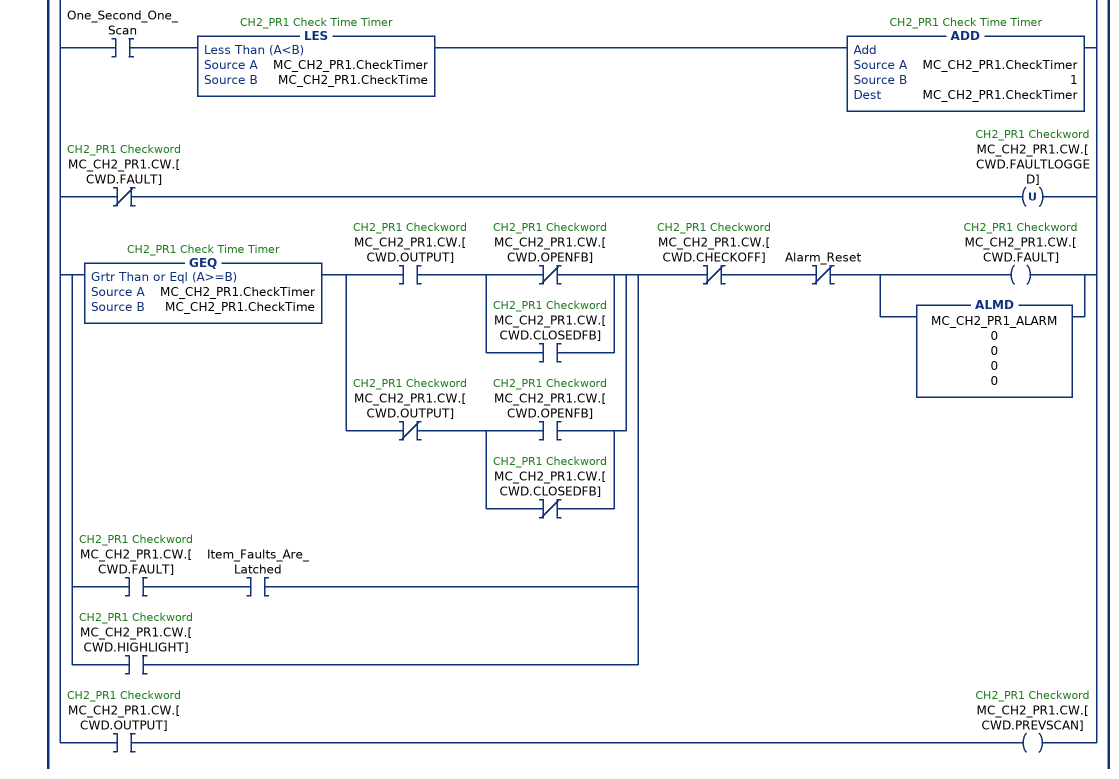
   38: [NEQ(MC_CH2_PR1.DriveBits,0) OTE(MC_CH2_PR1.CW.[CWD.AUTODRV]) ,[XIC(MC_CH2_PR1.CW.[CWD.AUTODRV]) XIO(MC_CH2_PR1.CW.[CWD.MANUAL]) ,XIC(MC_CH2_PR1.CW.[CWD.MANDRV]) XIC(MC_CH2_PR1.CW.[CWD.MANUAL]) ] OTE(MC_CH2_PR1.CW.[CWD.OUTPUT]) ,XIC(MC_CH2_PR1.CW.[CWD.OUTPUT]) OTE(MC_CH2_PR1_DR) ,XIC(S:FS) [OTU(MC_CH2_PR1.CW.[CWD.MANUAL]) ,LEQ(MC_CH2_PR1.CheckTime,0) MOV(Default_Check_Time,MC_CH2_PR1.CheckTime) ] ,[[XIC(MC_CH2_PR1_O) XIO(Item_Simulation_Flag) ,XIC(Item_Simulation_Flag) XIC(MC_CH2_PR1.CW.[CWD.OUTPUT]) XIO(MC_CH2_PR1.CW.[CWD.SIMFAIL]) ] OTE(MC_CH2_PR1.CW.[CWD.OPENFB]) ,[XIC(MC_CH2_PR1_C) XIO(Item_Simulation_Flag) ,XIC(Item_Simulation_Flag) XIO(MC_CH2_PR1.CW.[CWD.OUTPUT]) XIO(MC_CH2_PR1.CW.[CWD.SIMFAIL]) ] OTE(MC_CH2_PR1.CW.[CWD.CLOSEDFB]) ] ,[XIC(MC_CH2_PR1.CW.[CWD.OUTPUT]) XIO(MC_CH2_PR1.CW.[CWD.PREVSCAN]) ,XIO(MC_CH2_PR1.CW.[CWD.OUTPUT]) XIC(MC_CH2_PR1.CW.[CWD.PREVSCAN]) ] CLR(MC_CH2_PR1.CheckTimer) ,XIC(One_Second_One_Scan) LES(MC_CH2_PR1.CheckTimer,MC_CH2_PR1.CheckTime) ADD(MC_CH2_PR1.CheckTimer,1,MC_CH2_PR1.CheckTimer) ,XIO(MC_CH2_PR1.CW.[CWD.FAULT]) OTU(MC_CH2_PR1.CW.[CWD.FAULTLOGGED]) ,[GEQ(MC_CH2_PR1.CheckTimer,MC_CH2_PR1.CheckTime) [XIC(MC_CH2_PR1.CW.[CWD.OUTPUT]) [XIO(MC_CH2_PR1.CW.[CWD.OPENFB]) ,XIC(MC_CH2_PR1.CW.[CWD.CLOSEDFB]) ] ,XIO(MC_CH2_PR1.CW.[CWD.OUTPUT]) [XIC(MC_CH2_PR1.CW.[CWD.OPENFB]) ,XIO(MC_CH2_PR1.CW.[CWD.CLOSEDFB]) ] ] ,XIC(MC_CH2_PR1.CW.[CWD.FAULT]) XIC(Item_Faults_Are_Latched) ,XIC(MC_CH2_PR1.CW.[CWD.HIGHLIGHT]) ] XIO(MC_CH2_PR1.CW.[CWD.CHECKOFF]) XIO(Alarm_Reset) [OTE(MC_CH2_PR1.CW.[CWD.FAULT]) ,ALMD(MC_CH2_PR1_ALARM,0,0,0,0) ] ,XIC(MC_CH2_PR1.CW.[CWD.OUTPUT]) OTE(MC_CH2_PR1.CW.[CWD.PREVSCAN]) ];
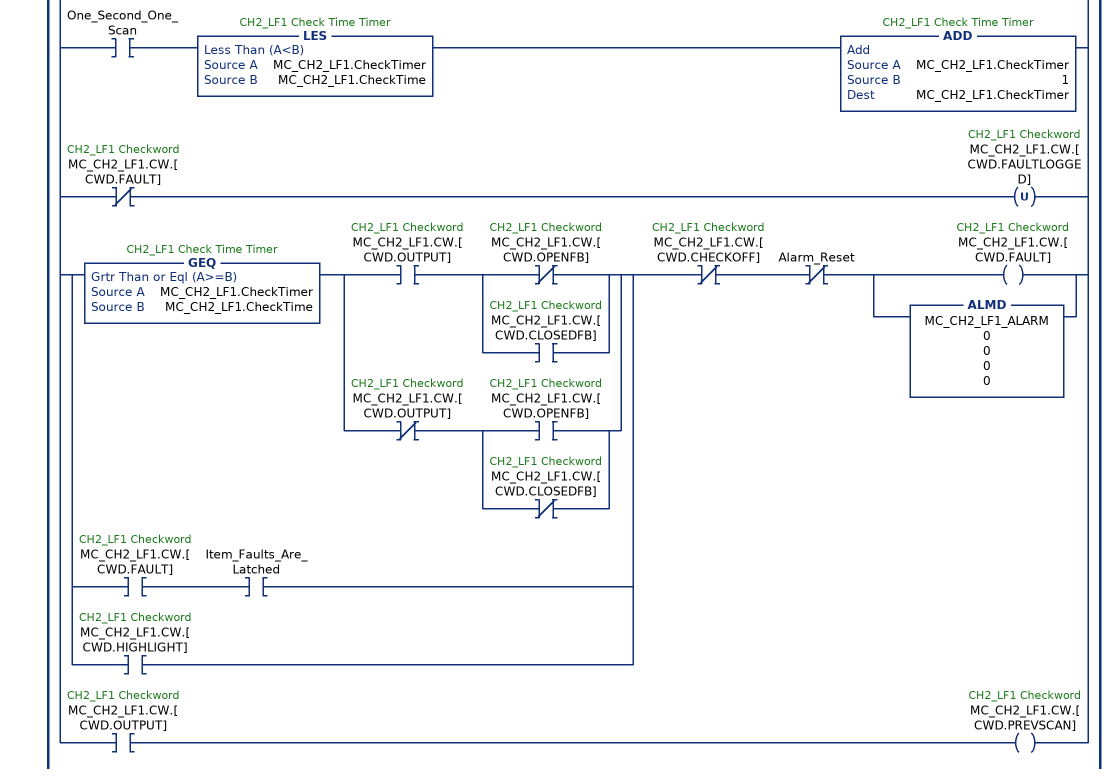
   39: [NEQ(MC_CH2_LF1.DriveBits,0) OTE(MC_CH2_LF1.CW.[CWD.AUTODRV]) ,[XIC(MC_CH2_LF1.CW.[CWD.AUTODRV]) XIO(MC_CH2_LF1.CW.[CWD.MANUAL]) ,XIC(MC_CH2_LF1.CW.[CWD.MANDRV]) XIC(MC_CH2_LF1.CW.[CWD.MANUAL]) ] OTE(MC_CH2_LF1.CW.[CWD.OUTPUT]) ,XIC(MC_CH2_LF1.CW.[CWD.OUTPUT]) OTE(MC_CH2_LF1_DR) ,XIC(S:FS) [OTU(MC_CH2_LF1.CW.[CWD.MANUAL]) ,LEQ(MC_CH2_LF1.CheckTime,0) MOV(Default_Check_Time,MC_CH2_LF1.CheckTime) ] ,[[XIC(MC_CH2_LF1_O) XIO(Item_Simulation_Flag) ,XIC(Item_Simulation_Flag) XIC(MC_CH2_LF1.CW.[CWD.OUTPUT]) XIO(MC_CH2_LF1.CW.[CWD.SIMFAIL]) ] OTE(MC_CH2_LF1.CW.[CWD.OPENFB]) ,[XIC(MC_CH2_LF1_C) XIO(Item_Simulation_Flag) ,XIC(Item_Simulation_Flag) XIO(MC_CH2_LF1.CW.[CWD.OUTPUT]) XIO(MC_CH2_LF1.CW.[CWD.SIMFAIL]) ] OTE(MC_CH2_LF1.CW.[CWD.CLOSEDFB]) ] ,[XIC(MC_CH2_LF1.CW.[CWD.OUTPUT]) XIO(MC_CH2_LF1.CW.[CWD.PREVSCAN]) ,XIO(MC_CH2_LF1.CW.[CWD.OUTPUT]) XIC(MC_CH2_LF1.CW.[CWD.PREVSCAN]) ] CLR(MC_CH2_LF1.CheckTimer) ,XIC(One_Second_One_Scan) LES(MC_CH2_LF1.CheckTimer,MC_CH2_LF1.CheckTime) ADD(MC_CH2_LF1.CheckTimer,1,MC_CH2_LF1.CheckTimer) ,XIO(MC_CH2_LF1.CW.[CWD.FAULT]) OTU(MC_CH2_LF1.CW.[CWD.FAULTLOGGED]) ,[GEQ(MC_CH2_LF1.CheckTimer,MC_CH2_LF1.CheckTime) [XIC(MC_CH2_LF1.CW.[CWD.OUTPUT]) [XIO(MC_CH2_LF1.CW.[CWD.OPENFB]) ,XIC(MC_CH2_LF1.CW.[CWD.CLOSEDFB]) ] ,XIO(MC_CH2_LF1.CW.[CWD.OUTPUT]) [XIC(MC_CH2_LF1.CW.[CWD.OPENFB]) ,XIO(MC_CH2_LF1.CW.[CWD.CLOSEDFB]) ] ] ,XIC(MC_CH2_LF1.CW.[CWD.FAULT]) XIC(Item_Faults_Are_Latched) ,XIC(MC_CH2_LF1.CW.[CWD.HIGHLIGHT]) ] XIO(MC_CH2_LF1.CW.[CWD.CHECKOFF]) XIO(Alarm_Reset) [OTE(MC_CH2_LF1.CW.[CWD.FAULT]) ,ALMD(MC_CH2_LF1_ALARM,0,0,0,0) ] ,XIC(MC_CH2_LF1.CW.[CWD.OUTPUT]) OTE(MC_CH2_LF1.CW.[CWD.PREVSCAN]) ];
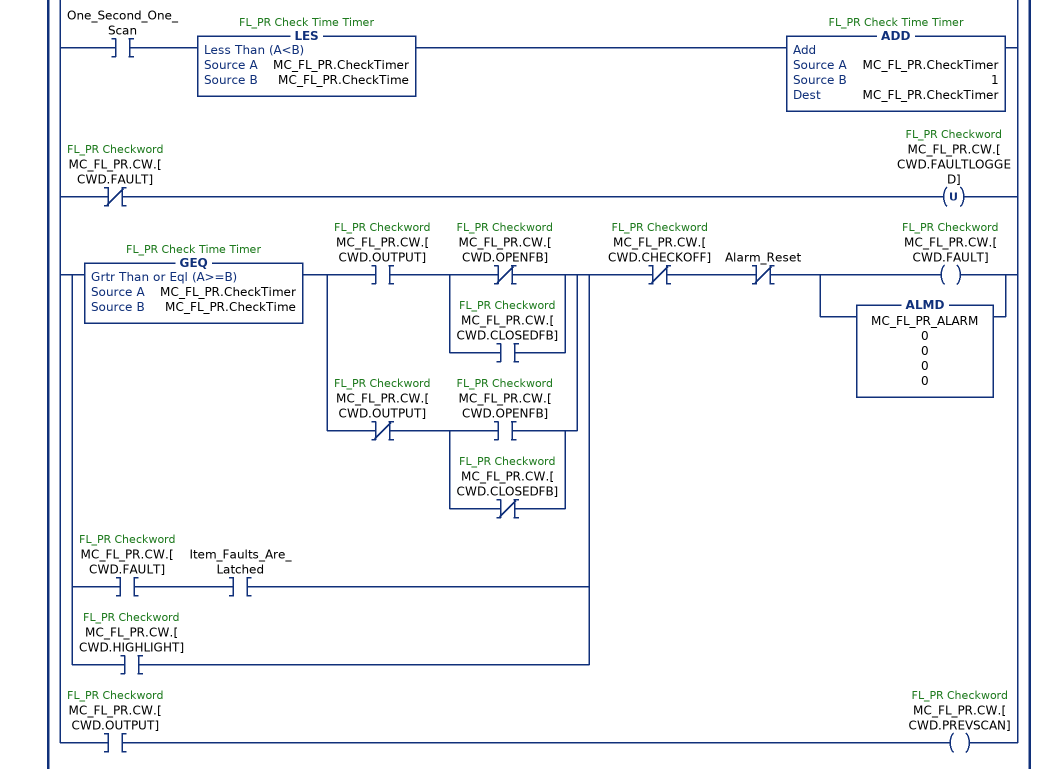
   40: [NEQ(MC_FL_PR.DriveBits,0) OTE(MC_FL_PR.CW.[CWD.AUTODRV]) ,[XIC(MC_FL_PR.CW.[CWD.AUTODRV]) XIO(MC_FL_PR.CW.[CWD.MANUAL]) ,XIC(MC_FL_PR.CW.[CWD.MANDRV]) XIC(MC_FL_PR.CW.[CWD.MANUAL]) ] OTE(MC_FL_PR.CW.[CWD.OUTPUT]) ,XIC(MC_FL_PR.CW.[CWD.OUTPUT]) OTE(MC_FL_PR_DR) ,XIC(S:FS) [OTU(MC_FL_PR.CW.[CWD.MANUAL]) ,LEQ(MC_FL_PR.CheckTime,0) MOV(Default_Check_Time,MC_FL_PR.CheckTime) ] ,[[XIC(MC_FL_PR_O) XIO(Item_Simulation_Flag) ,XIC(Item_Simulation_Flag) XIC(MC_FL_PR.CW.[CWD.OUTPUT]) XIO(MC_FL_PR.CW.[CWD.SIMFAIL]) ] OTE(MC_FL_PR.CW.[CWD.OPENFB]) ,[XIC(MC_FL_PR_C) XIO(Item_Simulation_Flag) ,XIC(Item_Simulation_Flag) XIO(MC_FL_PR.CW.[CWD.OUTPUT]) XIO(MC_FL_PR.CW.[CWD.SIMFAIL]) ] OTE(MC_FL_PR.CW.[CWD.CLOSEDFB]) ] ,[XIC(MC_FL_PR.CW.[CWD.OUTPUT]) XIO(MC_FL_PR.CW.[CWD.PREVSCAN]) ,XIO(MC_FL_PR.CW.[CWD.OUTPUT]) XIC(MC_FL_PR.CW.[CWD.PREVSCAN]) ] CLR(MC_FL_PR.CheckTimer) ,XIC(One_Second_One_Scan) LES(MC_FL_PR.CheckTimer,MC_FL_PR.CheckTime) ADD(MC_FL_PR.CheckTimer,1,MC_FL_PR.CheckTimer) ,XIO(MC_FL_PR.CW.[CWD.FAULT]) OTU(MC_FL_PR.CW.[CWD.FAULTLOGGED]) ,[GEQ(MC_FL_PR.CheckTimer,MC_FL_PR.CheckTime) [XIC(MC_FL_PR.CW.[CWD.OUTPUT]) [XIO(MC_FL_PR.CW.[CWD.OPENFB]) ,XIC(MC_FL_PR.CW.[CWD.CLOSEDFB]) ] ,XIO(MC_FL_PR.CW.[CWD.OUTPUT]) [XIC(MC_FL_PR.CW.[CWD.OPENFB]) ,XIO(MC_FL_PR.CW.[CWD.CLOSEDFB]) ] ] ,XIC(MC_FL_PR.CW.[CWD.FAULT]) XIC(Item_Faults_Are_Latched) ,XIC(MC_FL_PR.CW.[CWD.HIGHLIGHT]) ] XIO(MC_FL_PR.CW.[CWD.CHECKOFF]) XIO(Alarm_Reset) [OTE(MC_FL_PR.CW.[CWD.FAULT]) ,ALMD(MC_FL_PR_ALARM,0,0,0,0) ] ,XIC(MC_FL_PR.CW.[CWD.OUTPUT]) OTE(MC_FL_PR.CW.[CWD.PREVSCAN]) ];
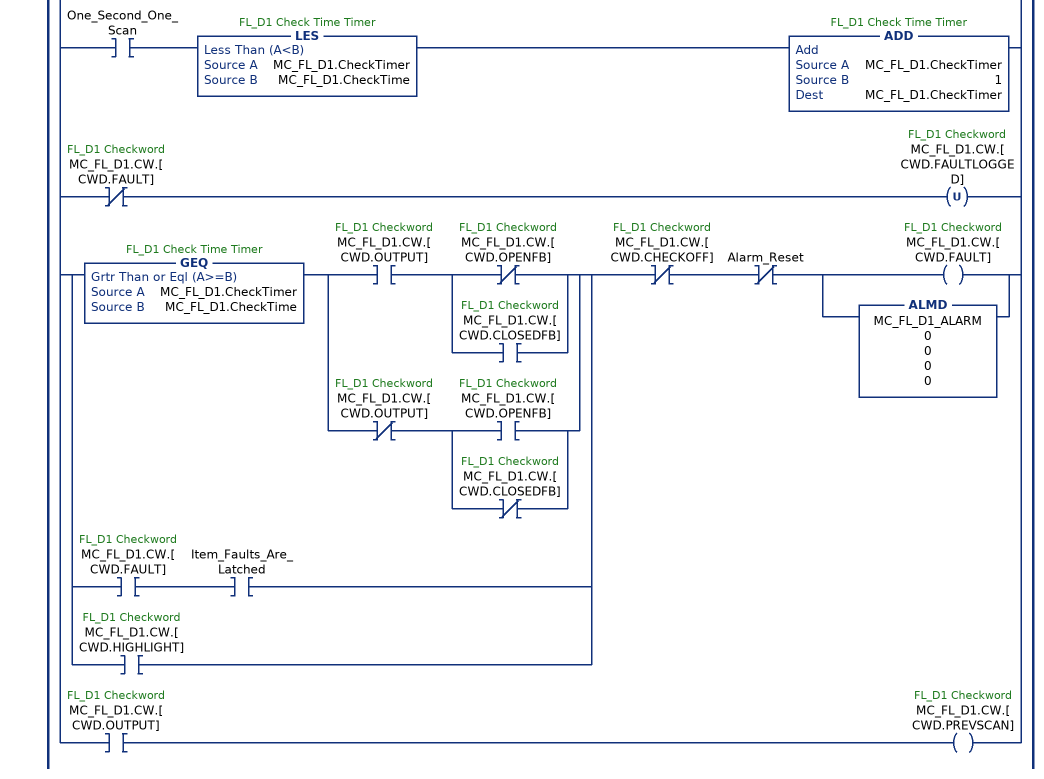
   41: [NEQ(MC_FL_D1.DriveBits,0) OTE(MC_FL_D1.CW.[CWD.AUTODRV]) ,[XIC(MC_FL_D1.CW.[CWD.AUTODRV]) XIO(MC_FL_D1.CW.[CWD.MANUAL]) ,XIC(MC_FL_D1.CW.[CWD.MANDRV]) XIC(MC_FL_D1.CW.[CWD.MANUAL]) ] OTE(MC_FL_D1.CW.[CWD.OUTPUT]) ,XIC(MC_FL_D1.CW.[CWD.OUTPUT]) OTE(MC_FL_D1_DR) ,XIC(S:FS) [OTU(MC_FL_D1.CW.[CWD.MANUAL]) ,LEQ(MC_FL_D1.CheckTime,0) MOV(Default_Check_Time,MC_FL_D1.CheckTime) ] ,[[XIC(MC_FL_D1_O) XIO(Item_Simulation_Flag) ,XIC(Item_Simulation_Flag) XIC(MC_FL_D1.CW.[CWD.OUTPUT]) XIO(MC_FL_D1.CW.[CWD.SIMFAIL]) ] OTE(MC_FL_D1.CW.[CWD.OPENFB]) ,[XIC(MC_FL_D1_C) XIO(Item_Simulation_Flag) ,XIC(Item_Simulation_Flag) XIO(MC_FL_D1.CW.[CWD.OUTPUT]) XIO(MC_FL_D1.CW.[CWD.SIMFAIL]) ] OTE(MC_FL_D1.CW.[CWD.CLOSEDFB]) ] ,[XIC(MC_FL_D1.CW.[CWD.OUTPUT]) XIO(MC_FL_D1.CW.[CWD.PREVSCAN]) ,XIO(MC_FL_D1.CW.[CWD.OUTPUT]) XIC(MC_FL_D1.CW.[CWD.PREVSCAN]) ] CLR(MC_FL_D1.CheckTimer) ,XIC(One_Second_One_Scan) LES(MC_FL_D1.CheckTimer,MC_FL_D1.CheckTime) ADD(MC_FL_D1.CheckTimer,1,MC_FL_D1.CheckTimer) ,XIO(MC_FL_D1.CW.[CWD.FAULT]) OTU(MC_FL_D1.CW.[CWD.FAULTLOGGED]) ,[GEQ(MC_FL_D1.CheckTimer,MC_FL_D1.CheckTime) [XIC(MC_FL_D1.CW.[CWD.OUTPUT]) [XIO(MC_FL_D1.CW.[CWD.OPENFB]) ,XIC(MC_FL_D1.CW.[CWD.CLOSEDFB]) ] ,XIO(MC_FL_D1.CW.[CWD.OUTPUT]) [XIC(MC_FL_D1.CW.[CWD.OPENFB]) ,XIO(MC_FL_D1.CW.[CWD.CLOSEDFB]) ] ] ,XIC(MC_FL_D1.CW.[CWD.FAULT]) XIC(Item_Faults_Are_Latched) ,XIC(MC_FL_D1.CW.[CWD.HIGHLIGHT]) ] XIO(MC_FL_D1.CW.[CWD.CHECKOFF]) XIO(Alarm_Reset) [OTE(MC_FL_D1.CW.[CWD.FAULT]) ,ALMD(MC_FL_D1_ALARM,0,0,0,0) ] ,XIC(MC_FL_D1.CW.[CWD.OUTPUT]) OTE(MC_FL_D1.CW.[CWD.PREVSCAN]) ];
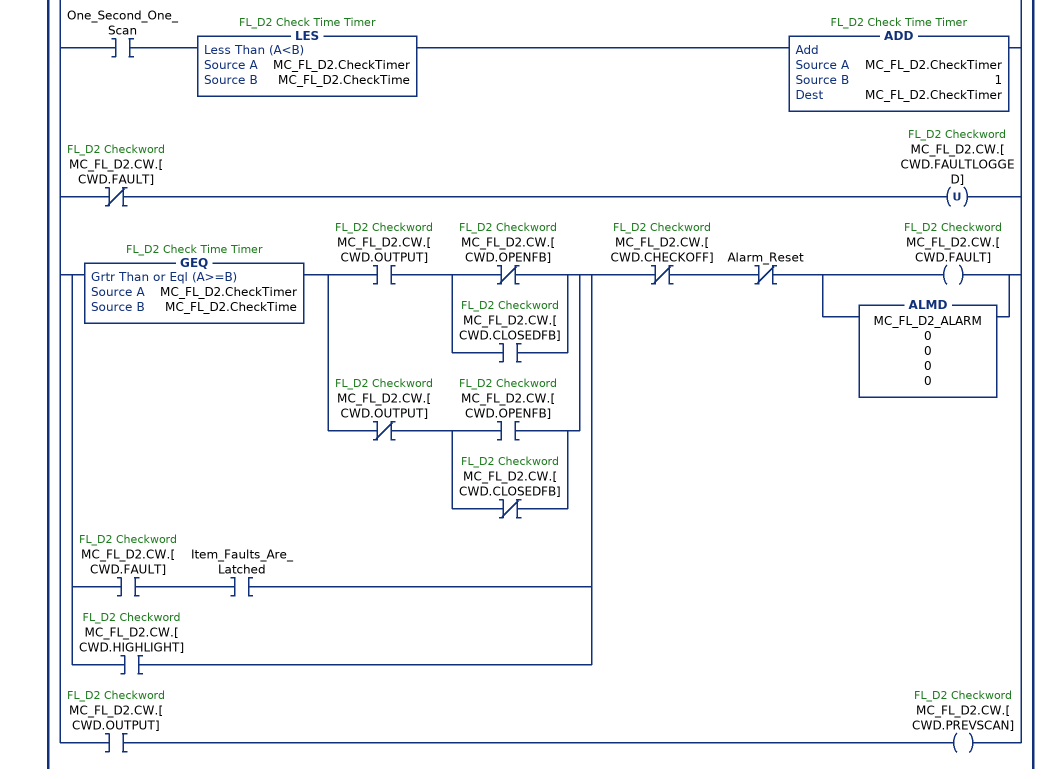
   42: [NEQ(MC_FL_D2.DriveBits,0) OTE(MC_FL_D2.CW.[CWD.AUTODRV]) ,[XIC(MC_FL_D2.CW.[CWD.AUTODRV]) XIO(MC_FL_D2.CW.[CWD.MANUAL]) ,XIC(MC_FL_D2.CW.[CWD.MANDRV]) XIC(MC_FL_D2.CW.[CWD.MANUAL]) ] OTE(MC_FL_D2.CW.[CWD.OUTPUT]) ,XIC(MC_FL_D2.CW.[CWD.OUTPUT]) OTE(MC_FL_D2_DR) ,XIC(S:FS) [OTU(MC_FL_D2.CW.[CWD.MANUAL]) ,LEQ(MC_FL_D2.CheckTime,0) MOV(Default_Check_Time,MC_FL_D2.CheckTime) ] ,[[XIC(MC_FL_D2_O) XIO(Item_Simulation_Flag) ,XIC(Item_Simulation_Flag) XIC(MC_FL_D2.CW.[CWD.OUTPUT]) XIO(MC_FL_D2.CW.[CWD.SIMFAIL]) ] OTE(MC_FL_D2.CW.[CWD.OPENFB]) ,[XIC(MC_FL_D2_C) XIO(Item_Simulation_Flag) ,XIC(Item_Simulation_Flag) XIO(MC_FL_D2.CW.[CWD.OUTPUT]) XIO(MC_FL_D2.CW.[CWD.SIMFAIL]) ] OTE(MC_FL_D2.CW.[CWD.CLOSEDFB]) ] ,[XIC(MC_FL_D2.CW.[CWD.OUTPUT]) XIO(MC_FL_D2.CW.[CWD.PREVSCAN]) ,XIO(MC_FL_D2.CW.[CWD.OUTPUT]) XIC(MC_FL_D2.CW.[CWD.PREVSCAN]) ] CLR(MC_FL_D2.CheckTimer) ,XIC(One_Second_One_Scan) LES(MC_FL_D2.CheckTimer,MC_FL_D2.CheckTime) ADD(MC_FL_D2.CheckTimer,1,MC_FL_D2.CheckTimer) ,XIO(MC_FL_D2.CW.[CWD.FAULT]) OTU(MC_FL_D2.CW.[CWD.FAULTLOGGED]) ,[GEQ(MC_FL_D2.CheckTimer,MC_FL_D2.CheckTime) [XIC(MC_FL_D2.CW.[CWD.OUTPUT]) [XIO(MC_FL_D2.CW.[CWD.OPENFB]) ,XIC(MC_FL_D2.CW.[CWD.CLOSEDFB]) ] ,XIO(MC_FL_D2.CW.[CWD.OUTPUT]) [XIC(MC_FL_D2.CW.[CWD.OPENFB]) ,XIO(MC_FL_D2.CW.[CWD.CLOSEDFB]) ] ] ,XIC(MC_FL_D2.CW.[CWD.FAULT]) XIC(Item_Faults_Are_Latched) ,XIC(MC_FL_D2.CW.[CWD.HIGHLIGHT]) ] XIO(MC_FL_D2.CW.[CWD.CHECKOFF]) XIO(Alarm_Reset) [OTE(MC_FL_D2.CW.[CWD.FAULT]) ,ALMD(MC_FL_D2_ALARM,0,0,0,0) ] ,XIC(MC_FL_D2.CW.[CWD.OUTPUT]) OTE(MC_FL_D2.CW.[CWD.PREVSCAN]) ];
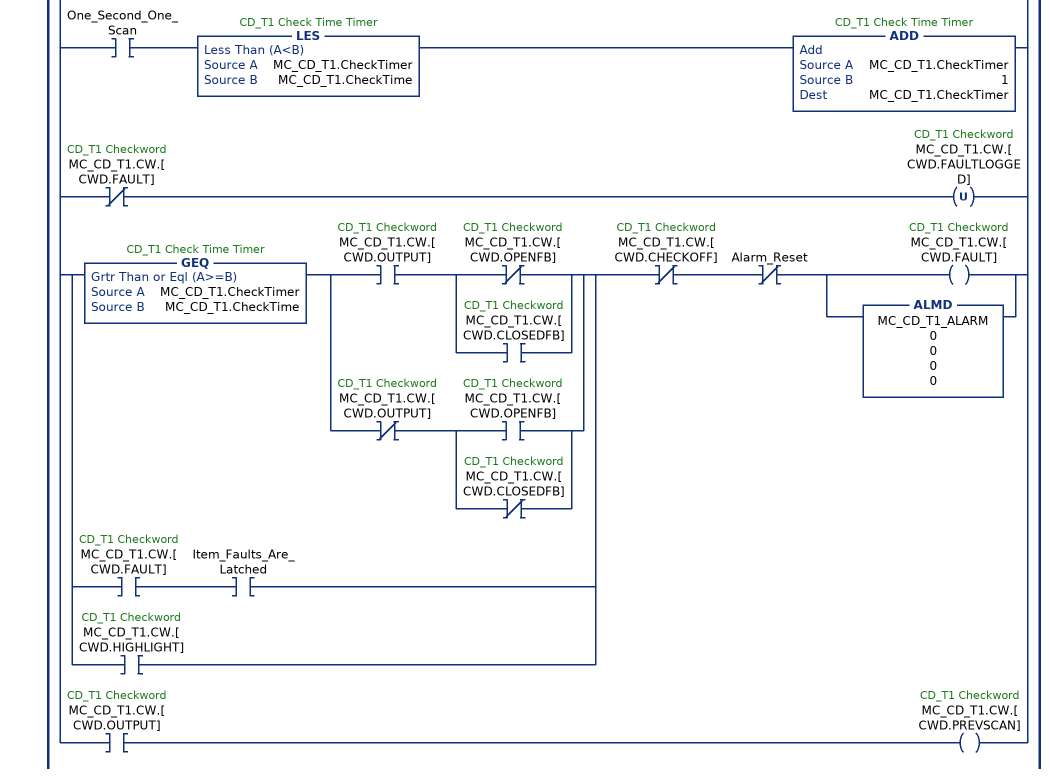
   43: [NEQ(MC_CD_T1.DriveBits,0) OTE(MC_CD_T1.CW.[CWD.AUTODRV]) ,[XIC(MC_CD_T1.CW.[CWD.AUTODRV]) XIO(MC_CD_T1.CW.[CWD.MANUAL]) ,XIC(MC_CD_T1.CW.[CWD.MANDRV]) XIC(MC_CD_T1.CW.[CWD.MANUAL]) ] OTE(MC_CD_T1.CW.[CWD.OUTPUT]) ,XIC(MC_CD_T1.CW.[CWD.OUTPUT]) OTE(MC_CD_T1_DR) ,XIC(S:FS) [OTU(MC_CD_T1.CW.[CWD.MANUAL]) ,LEQ(MC_CD_T1.CheckTime,0) MOV(Default_Check_Time,MC_CD_T1.CheckTime) ] ,[[XIC(MC_CD_T1_O) XIO(Item_Simulation_Flag) ,XIC(Item_Simulation_Flag) XIC(MC_CD_T1.CW.[CWD.OUTPUT]) XIO(MC_CD_T1.CW.[CWD.SIMFAIL]) ] OTE(MC_CD_T1.CW.[CWD.OPENFB]) ,[XIC(MC_CD_T1_C) XIO(Item_Simulation_Flag) ,XIC(Item_Simulation_Flag) XIO(MC_CD_T1.CW.[CWD.OUTPUT]) XIO(MC_CD_T1.CW.[CWD.SIMFAIL]) ] OTE(MC_CD_T1.CW.[CWD.CLOSEDFB]) ] ,[XIC(MC_CD_T1.CW.[CWD.OUTPUT]) XIO(MC_CD_T1.CW.[CWD.PREVSCAN]) ,XIO(MC_CD_T1.CW.[CWD.OUTPUT]) XIC(MC_CD_T1.CW.[CWD.PREVSCAN]) ] CLR(MC_CD_T1.CheckTimer) ,XIC(One_Second_One_Scan) LES(MC_CD_T1.CheckTimer,MC_CD_T1.CheckTime) ADD(MC_CD_T1.CheckTimer,1,MC_CD_T1.CheckTimer) ,XIO(MC_CD_T1.CW.[CWD.FAULT]) OTU(MC_CD_T1.CW.[CWD.FAULTLOGGED]) ,[GEQ(MC_CD_T1.CheckTimer,MC_CD_T1.CheckTime) [XIC(MC_CD_T1.CW.[CWD.OUTPUT]) [XIO(MC_CD_T1.CW.[CWD.OPENFB]) ,XIC(MC_CD_T1.CW.[CWD.CLOSEDFB]) ] ,XIO(MC_CD_T1.CW.[CWD.OUTPUT]) [XIC(MC_CD_T1.CW.[CWD.OPENFB]) ,XIO(MC_CD_T1.CW.[CWD.CLOSEDFB]) ] ] ,XIC(MC_CD_T1.CW.[CWD.FAULT]) XIC(Item_Faults_Are_Latched) ,XIC(MC_CD_T1.CW.[CWD.HIGHLIGHT]) ] XIO(MC_CD_T1.CW.[CWD.CHECKOFF]) XIO(Alarm_Reset) [OTE(MC_CD_T1.CW.[CWD.FAULT]) ,ALMD(MC_CD_T1_ALARM,0,0,0,0) ] ,XIC(MC_CD_T1.CW.[CWD.OUTPUT]) OTE(MC_CD_T1.CW.[CWD.PREVSCAN]) ];
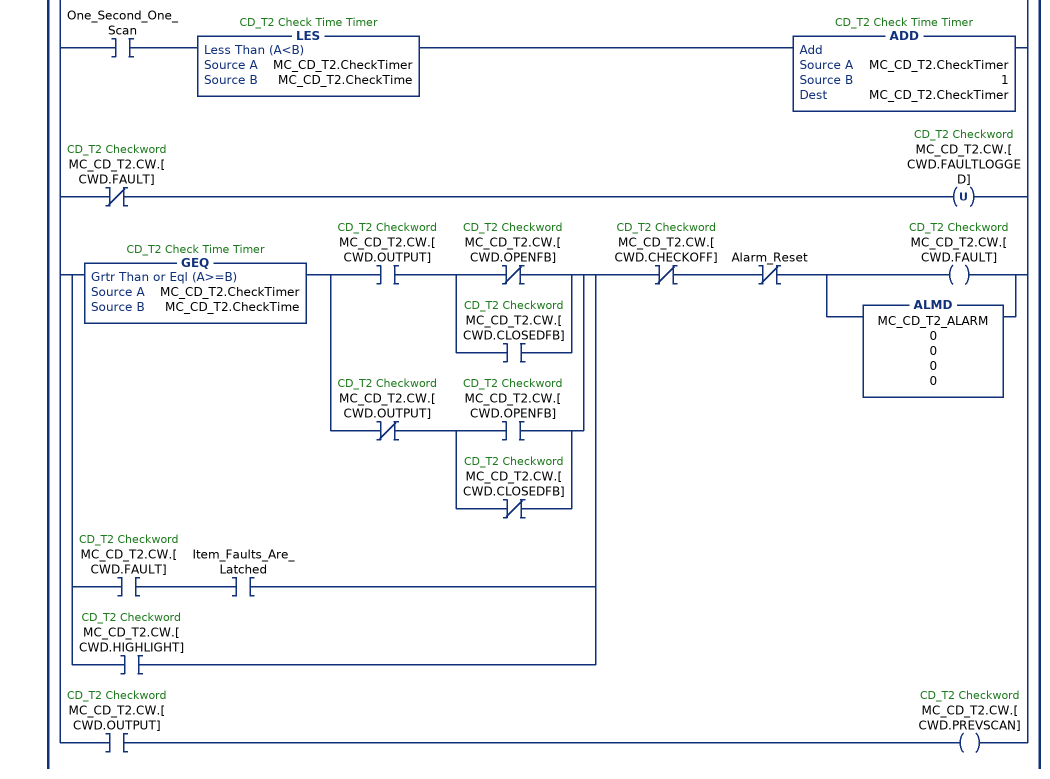
   44: [NEQ(MC_CD_T2.DriveBits,0) OTE(MC_CD_T2.CW.[CWD.AUTODRV]) ,[XIC(MC_CD_T2.CW.[CWD.AUTODRV]) XIO(MC_CD_T2.CW.[CWD.MANUAL]) ,XIC(MC_CD_T2.CW.[CWD.MANDRV]) XIC(MC_CD_T2.CW.[CWD.MANUAL]) ] OTE(MC_CD_T2.CW.[CWD.OUTPUT]) ,XIC(MC_CD_T2.CW.[CWD.OUTPUT]) OTE(MC_CD_T2_DR) ,XIC(S:FS) [OTU(MC_CD_T2.CW.[CWD.MANUAL]) ,LEQ(MC_CD_T2.CheckTime,0) MOV(Default_Check_Time,MC_CD_T2.CheckTime) ] ,[[XIC(MC_CD_T2_O) XIO(Item_Simulation_Flag) ,XIC(Item_Simulation_Flag) XIC(MC_CD_T2.CW.[CWD.OUTPUT]) XIO(MC_CD_T2.CW.[CWD.SIMFAIL]) ] OTE(MC_CD_T2.CW.[CWD.OPENFB]) ,[XIC(MC_CD_T2_C) XIO(Item_Simulation_Flag) ,XIC(Item_Simulation_Flag) XIO(MC_CD_T2.CW.[CWD.OUTPUT]) XIO(MC_CD_T2.CW.[CWD.SIMFAIL]) ] OTE(MC_CD_T2.CW.[CWD.CLOSEDFB]) ] ,[XIC(MC_CD_T2.CW.[CWD.OUTPUT]) XIO(MC_CD_T2.CW.[CWD.PREVSCAN]) ,XIO(MC_CD_T2.CW.[CWD.OUTPUT]) XIC(MC_CD_T2.CW.[CWD.PREVSCAN]) ] CLR(MC_CD_T2.CheckTimer) ,XIC(One_Second_One_Scan) LES(MC_CD_T2.CheckTimer,MC_CD_T2.CheckTime) ADD(MC_CD_T2.CheckTimer,1,MC_CD_T2.CheckTimer) ,XIO(MC_CD_T2.CW.[CWD.FAULT]) OTU(MC_CD_T2.CW.[CWD.FAULTLOGGED]) ,[GEQ(MC_CD_T2.CheckTimer,MC_CD_T2.CheckTime) [XIC(MC_CD_T2.CW.[CWD.OUTPUT]) [XIO(MC_CD_T2.CW.[CWD.OPENFB]) ,XIC(MC_CD_T2.CW.[CWD.CLOSEDFB]) ] ,XIO(MC_CD_T2.CW.[CWD.OUTPUT]) [XIC(MC_CD_T2.CW.[CWD.OPENFB]) ,XIO(MC_CD_T2.CW.[CWD.CLOSEDFB]) ] ] ,XIC(MC_CD_T2.CW.[CWD.FAULT]) XIC(Item_Faults_Are_Latched) ,XIC(MC_CD_T2.CW.[CWD.HIGHLIGHT]) ] XIO(MC_CD_T2.CW.[CWD.CHECKOFF]) XIO(Alarm_Reset) [OTE(MC_CD_T2.CW.[CWD.FAULT]) ,ALMD(MC_CD_T2_ALARM,0,0,0,0) ] ,XIC(MC_CD_T2.CW.[CWD.OUTPUT]) OTE(MC_CD_T2.CW.[CWD.PREVSCAN]) ];
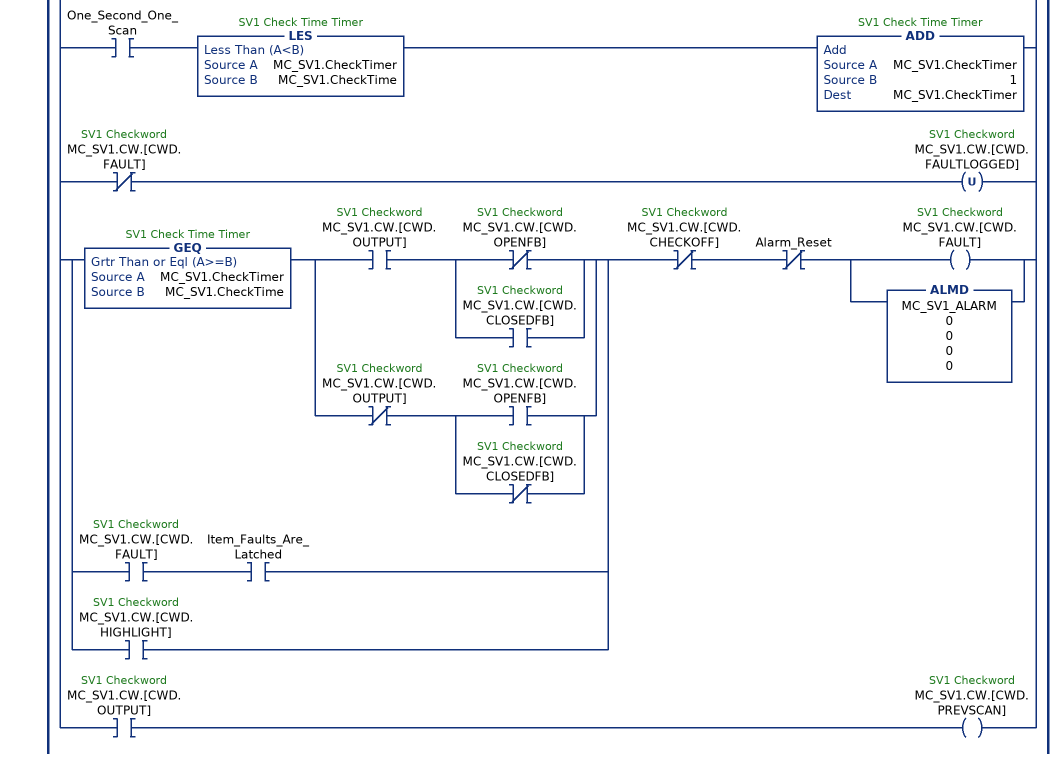
   45: [NEQ(MC_SV1.DriveBits,0) OTE(MC_SV1.CW.[CWD.AUTODRV]) ,[XIC(MC_SV1.CW.[CWD.AUTODRV]) XIO(MC_SV1.CW.[CWD.MANUAL]) ,XIC(MC_SV1.CW.[CWD.MANDRV]) XIC(MC_SV1.CW.[CWD.MANUAL]) ] OTE(MC_SV1.CW.[CWD.OUTPUT]) ,XIC(MC_SV1.CW.[CWD.OUTPUT]) OTE(MC_SV1_DR) ,XIC(S:FS) [OTU(MC_SV1.CW.[CWD.MANUAL]) ,LEQ(MC_SV1.CheckTime,0) MOV(Default_Check_Time,MC_SV1.CheckTime) ] ,[[XIC(MC_SV1_O) XIO(Item_Simulation_Flag) ,XIC(Item_Simulation_Flag) XIC(MC_SV1.CW.[CWD.OUTPUT]) XIO(MC_SV1.CW.[CWD.SIMFAIL]) ] OTE(MC_SV1.CW.[CWD.OPENFB]) ,[XIC(MC_SV1_C) XIO(Item_Simulation_Flag) ,XIC(Item_Simulation_Flag) XIO(MC_SV1.CW.[CWD.OUTPUT]) XIO(MC_SV1.CW.[CWD.SIMFAIL]) ] OTE(MC_SV1.CW.[CWD.CLOSEDFB]) ] ,[XIC(MC_SV1.CW.[CWD.OUTPUT]) XIO(MC_SV1.CW.[CWD.PREVSCAN]) ,XIO(MC_SV1.CW.[CWD.OUTPUT]) XIC(MC_SV1.CW.[CWD.PREVSCAN]) ] CLR(MC_SV1.CheckTimer) ,XIC(One_Second_One_Scan) LES(MC_SV1.CheckTimer,MC_SV1.CheckTime) ADD(MC_SV1.CheckTimer,1,MC_SV1.CheckTimer) ,XIO(MC_SV1.CW.[CWD.FAULT]) OTU(MC_SV1.CW.[CWD.FAULTLOGGED]) ,[GEQ(MC_SV1.CheckTimer,MC_SV1.CheckTime) [XIC(MC_SV1.CW.[CWD.OUTPUT]) [XIO(MC_SV1.CW.[CWD.OPENFB]) ,XIC(MC_SV1.CW.[CWD.CLOSEDFB]) ] ,XIO(MC_SV1.CW.[CWD.OUTPUT]) [XIC(MC_SV1.CW.[CWD.OPENFB]) ,XIO(MC_SV1.CW.[CWD.CLOSEDFB]) ] ] ,XIC(MC_SV1.CW.[CWD.FAULT]) XIC(Item_Faults_Are_Latched) ,XIC(MC_SV1.CW.[CWD.HIGHLIGHT]) ] XIO(MC_SV1.CW.[CWD.CHECKOFF]) XIO(Alarm_Reset) [OTE(MC_SV1.CW.[CWD.FAULT]) ,ALMD(MC_SV1_ALARM,0,0,0,0) ] ,XIC(MC_SV1.CW.[CWD.OUTPUT]) OTE(MC_SV1.CW.[CWD.PREVSCAN]) ];